
screen "设置画面" 1280x740, template "模板_设置"
   on GenerateScreen: "TitleUpdater"()
   TextField "Text Field_2" at 90,72 size 116x49; Text '总捻度:'
   TextField "Text Field_6" at 320,72 size 107x49; Text '捻/米'
   TextField "Text Field_19" at 674,70 size 140x49; Text '捻缩捻度:'
   TextField "Text Field_20" at 674,133 size 140x49; Text '捻缩距离:'
   TextField "Text Field_21" at 674,196 size 140x49; Text '捻缩时间:'
   TextField "Text Field_22" at 674,259 size 140x49; Text '捻缩速度:'
   TextField "Text Field_15" at 786,14 size 154x42; Text '捻缩设定'
   TextField "Text Field_29" at 753,476 size 140x49; Text '成纱支数:'
   TextField "Text Field_31" at 674,322 size 140x49; Text '卷绕长度:'
   TextField "Text Field_32" at 940,70 size 98x49; Text '捻/米'
   TextField "Text Field_33" at 940,133 size 98x49; Text 'mm'
   TextField "Text Field_34" at 940,196 size 98x49; Text '秒'
   TextField "Text Field_35" at 940,259 size 98x49; Text 'mm/s'
   TextField "Text Field_36" at 940,322 size 98x49; Text 'mm'
   TextField "Text Field_48" at 552,72 size 84x49; Text '秒'
   TextField "Text Field_40" at 791,420 size 228x42; Text '成形、张力设定'
   TextField "Text Field_41" at 753,539 size 140x49; Text '纱穗个数:'
   TextField "Text Field_41#mig1" at 753,602 size 140x49; Text '单纱张力:'
   TextField "Text Field_14" at 142,14 size 336x42; Text '捻度设定分配/锭速设定'
   TextField "Text Field_25" at 96,477 size 133x48; Text '总牵伸:'
   TextField "Text Field_26" at 96,540 size 133x49; Text '送条牵伸:'
   TextField "Text Field_1" at 365,420 size 193x42; Text '牵伸设定分配'
   TextField "Text Field_28" at 348,540 size 212x49; Text '第一牵伸(3段):'
   TextField "Text Field_37" at 348,603 size 212x49; Text '集中牵伸区(3段):'
   TextField "Text Field_38" at 348,477 size 212x48; Text '第一牵伸区(3段):'
   TextField "Text Field_39" at 666,477 size 32x48; Text 'mm'
   TextField "Text Field_42" at 666,603 size 32x49; Text 'mm'
   TextField "Text Field_27" at 43,603 size 186x49; Text '分散牵伸(2段):'
   SymbolicIOField "符号 IO 域_1" at 229,420 size 106x44; TextOn '1'; TextOff '0'; TextList "QainShen_Select"
      ProcessValue <- "ST_HMI_Var_HMI_i16_QianShen_Select"
   IOField "IO Field_14" at 229,477 size 106x48; FormatPattern 9.99
      ProcessValue <- "ST_HMI_Var_HMI_r64QianShen_All"
   IOField "IO Field_15" at 229,540 size 106x49; FormatPattern 9.999
      ProcessValue <- "ST_HMI_Var_HMI_r64QianShen_WuNian"
   IOField "IO Field_17" at 560,540 size 93x49; FormatPattern 9.99
      ProcessValue <- "ST_HMI_Var_HMI_r64QianShen_First"
   IOField "IO Field_20" at 560,603 size 93x49; FormatPattern 99
      ProcessValue <- "ST_HMI_Var_HMI_r64QianShen_finalArea"
   IOField "IO Field_21" at 560,477 size 93x48; FormatPattern 999
      ProcessValue <- "ST_HMI_Var_HMI_r64QianShen_FirstArea"
   IOField "IO Field_16" at 229,603 size 106x49; FormatPattern 9.99
      ProcessValue <- "ST_HMI_Var_HMI_r64QianShen_FenSan"
   TextField "Text Field_3" at 66,136 size 140x47; Text '牵伸捻度:'
   IOField "IO Field_1" at 208,136 size 104x49; FormatPattern 999
      on OnFinishInput: SetBit("ST_Calculation_Var_HMI_bo_Calculation_0_Start"); SetTag("ST_Calculation_Var_g_i16_Calculation_0_3_Select_Status", 1)
      ProcessValue <- "ST_HMI_Var_HMI_r64NianDu_QianShen_Best"
   TextField "Text Field_4" at 320,136 size 107x49; Text '捻/米'
   TextField "Text Field_5" at 552,136 size 84x49; Text '转/分'
   IOField "IO Field_3" at 208,200 size 104x49; FormatPattern 9.99
      on OnFinishInput: SetBit("ST_Calculation_Var_HMI_bo_Calculation_0_Start"); SetTag("ST_Calculation_Var_g_i16_Calculation_0_3_Select_Status", 1)
      ProcessValue <- "ST_HMI_Var_HMI_r64Ratio_PositiveAccel_Jerk_JiaNian"
   TextField "Text Field_8" at 66,264 size 140x47; Text '追捻:'
   Button "OBJECT_107" at 208,264 size 104x48; TextOff '启用 / EXIT'
      on Release: SetBit("ST_HMI_Var_HMI_boNianDu_3")
      on Change: SetBit("ST_Calculation_Var_HMI_bo_Calculation_0_Start"); SetTag("ST_Calculation_Var_g_i16_Calculation_0_3_Select_Status", 1)
      Appearance <- "ST_HMI_Var_HMI_boNianDu_3"
   Button "OBJECT_1" at 432,264 size 112x48; TextOff '停用 / EXIT'
      on Release: ResetBit("ST_HMI_Var_HMI_boNianDu_3")
      on Change: SetBit("ST_Calculation_Var_HMI_bo_Calculation_0_Start"); SetTag("ST_Calculation_Var_g_i16_Calculation_0_3_Select_Status", 1)
      Appearance <- "ST_HMI_Var_HMI_boNianDu_3"
   TextField "Text Field_9" at 24,328 size 182x47; Text '追捻开始捻度:'
   IOField "IO Field_4" at 208,328 size 104x49; FormatPattern 9999
      on OnFinishInput: SetBit("ST_Calculation_Var_HMI_bo_Calculation_0_Start"); SetTag("ST_Calculation_Var_g_i16_Calculation_0_3_Select_Status", 1)
      ProcessValue <- "ST_HMI_Var_HMI_r64NianDu_1"
   TextField "Text Field_10" at 328,328 size 84x49; Text '捻/米'
   TextField "Text Field_11" at 552,328 size 84x49; Text '转/分'
   TextField "Text Field_12" at 320,200 size 107x47; Text '加速度:'
   IOField "IO Field_5" at 432,328 size 112x49; FormatPattern 99999
      on OnFinishInput: SetBit("ST_Calculation_Var_HMI_bo_Calculation_0_Start"); SetTag("ST_Calculation_Var_g_i16_Calculation_0_3_Select_Status", 1)
      ProcessValue <- "ST_HMI_Var_HMI_r64NianSu_2"
   TextField "Text Field_7" at 48,202 size 158x47; Text '加速度比例:'
   IOField "IO Field_43" at 208,72 size 104x49; FormatPattern 9999
      on OnFinishInput: SetBit("ST_Calculation_Var_HMI_bo_Calculation_0_Start"); SetTag("ST_Calculation_Var_g_i16_Calculation_0_3_Select_Status", 1)
      ProcessValue <- "ST_HMI_Var_HMI_r64NianDu_all"
   IOField "IO Field_13" at 432,72 size 112x49; FormatPattern 99.9
      ProcessValue <- "ST_HMI_Var_HMI_r64Time_JiaNian"
      Appearance <- "ST_HMI_Var_HMI_boAlarm_NianDu_Time"
   IOField "IO Field_9" at 814,70 size 112x49; FormatPattern 9999
      on OnFinishInput: SetBit("ST_Calculation_Var_HMI_bo_Calculation_0_Start"); SetTag("ST_Calculation_Var_g_i16_Calculation_0_3_Select_Status", 1)
      ProcessValue <- "ST_HMI_Var_HMI_r64NianDu_NianSuo"
   IOField "IO Field_10" at 814,133 size 112x49; FormatPattern 999
      on OnFinishInput: SetBit("ST_Calculation_Var_HMI_bo_Calculation_0_Start")
      Appearance <- "ST_HMI_Var_HMI_boAlarm_NianSuo_PosNon"
      ProcessValue <- "ST_HMI_Var_HMI_r64Position_NianSuo"
   IOField "IO Field_11" at 814,196 size 112x49; FormatPattern 99.9
      ProcessValue <- "ST_HMI_Var_HMI_r64Time_NianSuo"
   IOField "IO Field_12" at 814,259 size 112x49; FormatPattern 99.9
      ProcessValue <- "ST_HMI_Var_HMI_r64Velocity_NianSuo"
      Appearance <- "ST_HMI_Var_HMI_boAlarm_NianSuo_SuDuOver"
   IOField "IO Field_19" at 814,322 size 112x49; FormatPattern 9999
      ProcessValue <- "ST_HMI_Var_HMI_r64Length_JuanRao"
   IOField "IO Field_18" at 907,476 size 126x49; FormatPattern 99.99
      ProcessValue <- "ST_HMI_Var_HMI_r64ZhiShu_ChengSha"
   IOField "IO Field_75" at 907,539 size 126x49; FormatPattern 9999
      ProcessValue <- "ST_HMI_Var_HMI_r64_ShuLiang_ShaSui"
   IOField "IO Field_76" at 907,602 size 126x49; FormatPattern 999.9
      ProcessValue <- "ST_HMI_Var_HMI_r64_LuoSha_Force_DanSha_ZhangLi_FangKai"
   IOField "IO Field_2" at 432,136 size 112x49; FormatPattern 99999
      ProcessValue <- "ST_HMI_Var_HMI_r64NianSu_Max"
      Appearance <- "ST_HMI_Var_HMI_boAlarm_NianDu_Time"
   IOField "IO Field_6" at 432,200 size 112x49; FormatPattern 99999
      Visibility <- "ST_Calculation_Var_Date_Temp"
      ProcessValue <- "ST_Calculation_Var_g_r64Axis_DingZi_PositiveAccel_Buffer_JiaNian{0}"
      Appearance <- "ST_HMI_Var_HMI_boAlarm_NianDu_Time"
   IOField "IO Field_8" at 432,200 size 112x49; FormatPattern 99999
      Visibility <- "ST_Calculation_Var_Date_Temp"
      ProcessValue <- "ST_Calculation_Var_g_r64Axis_DingZi_PositiveAccel_Buffer_JiaNian{1}"
      Appearance <- "ST_HMI_Var_HMI_boAlarm_NianDu_Time"
   TextField "文本域_5" at 1,304 size 880x170; Text '捻度报警！设置捻度为 ，实际捻度为 ， 已自动停止，请检查设置画面参数，重新设置总捻度， 检查设置其他参数，使画面上的参数没有红色闪烁，然 后按“启动”，若继续出现此报警，请从生头重新开始'
      Visibility <- "ST_HMI_Var_HMI_i16_NianduAlarmStatus"
   IOField "IO Field_7" at 322,305 size 86x32; FormatPattern 9999
      on OnFinishInput: SetBit("ST_Calculation_Var_HMI_bo_Calculation_0_Start"); SetTag("ST_Calculation_Var_g_i16_Calculation_0_3_Select_Status", 1)
      Visibility <- "ST_HMI_Var_HMI_i16_NianduAlarmStatus"
      ProcessValue <- "ST_HMI_Var_HMI_r64NianDu_all"
   IOField "IO Field_22" at 601,305 size 86x32; FormatPattern 9999
      Visibility <- "ST_HMI_Var_HMI_i16_NianduAlarmStatus"
      ProcessValue <- "ST_HMI_Var_HMI_r64Niandu_all_Current"
   Button "按钮_16" at 734,414 size 137x44; TextOff '知道了'
      on Click: SetTag("ST_HMI_Var_HMI_i16_NianduAlarmStatus", 0); SetBit("ST_Calculation_Var_HMI_bo_Calculation_0_Start"); ResetBit("ST_HMI_Var_HMI_bo_XiangLing")
      Visibility <- "ST_HMI_Var_HMI_i16_NianduAlarmStatus"
   Circle "圆_4" at 774,325 size 60x60
      Visibility <- "ST_HMI_Var_HMI_i16_NianduAlarmStatus"
      Appearance <- "ST_HMI_Var_HMI_bo_XiangLing"
   TextField "文本域_10" at 7,311 size 880x170; Text '锭子不转报警！请至报警画面解除报警，然后点击“退 出紧急停止”，点击“启动”开机，或者按正常步骤断电 重启，然后开机'
      Visibility <- "ST_HMI_Var_HMI_i16_Dingzi_50102AlarmStatus"
   Button "按钮_6" at 732,413 size 137x44; TextOff '知道了'
      on Click: SetTag("ST_HMI_Var_HMI_i16_Dingzi_50102AlarmStatus", 0); ResetBit("ST_HMI_Var_HMI_bo_XiangLing")
      Visibility <- "ST_HMI_Var_HMI_i16_Dingzi_50102AlarmStatus"
   Circle "圆_1" at 772,324 size 60x60
      Visibility <- "ST_HMI_Var_HMI_i16_Dingzi_50102AlarmStatus"
      Appearance <- "ST_HMI_Var_HMI_bo_XiangLing"

screen "时间显示" 1280x740, template "模板_根"
   on GenerateScreen: "TitleUpdater"(); "timeConverse"()
   Button "HmiScreenItemData_8" at 1120,65 size 159x47; TextOn '向后'; TextOff '向后'
      on Release: ActivateScreen("友联走架智控系统", 0)
   Button "按钮_1" at 174,88 size 95x82; TextOff '出车'
      Appearance <- "ST_Main_Var_g_i16_Automatic_Status"
   Button "按钮_2" at 321,88 size 95x82; TextOff '加捻'
      Appearance <- "ST_Main_Var_g_i16_Automatic_Status"
   Button "按钮_3" at 467,88 size 96x82; TextOff '退绕'
      Appearance <- "ST_Main_Var_g_i16_Automatic_Status"
   Button "按钮_4" at 614,88 size 95x82; TextOff '进车'
      Appearance <- "ST_Main_Var_g_i16_Automatic_Status"
   Button "按钮_5" at 760,88 size 96x82; TextOff '周期'
      Appearance <- "ST_Main_Var_g_i16_Automatic_Status"
   TextField "文本域_1" at 51,360 size 207x37; Text '系统总运行时间:'
   TextField "文本域_2" at 346,360 size 56x37; Text '年'
   TextField "文本域_4" at 460,360 size 56x37; Text '天'
   TextField "文本域_5" at 563,360 size 56x37; Text '时'
   TextField "文本域_6" at 661,360 size 56x37; Text '分'
   TextField "文本域_7" at 760,360 size 56x37; Text '秒'
   IOField "IO Field_23" at 174,183 size 95x55; FormatPattern 99.99
      ProcessValue <- "ST_Main_Var_g_r64_Time_chuche"
   IOField "IO Field_24" at 321,183 size 95x55; FormatPattern 99.99
      ProcessValue <- "ST_Main_Var_g_r64_Time_jianian"
   IOField "IO Field_25" at 467,183 size 96x55; FormatPattern 99.99
      ProcessValue <- "ST_Main_Var_g_r64_Time_tuirao"
   IOField "IO Field_26" at 614,183 size 95x55; FormatPattern 99.99
      ProcessValue <- "ST_Main_Var_g_r64_Time_juanrao"
   IOField "IO Field_27" at 760,183 size 96x55; FormatPattern 99.99
      ProcessValue <- "ST_Main_Var_g_r64_Time_Once"
   IOField "IO Field_29" at 269,350 size 72x55; FormatPattern 999
      ProcessValue <- "VBS_time_year"
   IOField "IO Field_30" at 385,350 size 68x55; FormatPattern 999
      ProcessValue <- "VBS_time_day"
   IOField "IO Field_30#mig1" at 499,350 size 55x55; FormatPattern 99
      ProcessValue <- "VBS_time_hour"
   IOField "IO Field_31" at 600,350 size 55x55; FormatPattern 99
      ProcessValue <- "VBS_time_min"
   IOField "IO Field_32" at 701,350 size 52x55; FormatPattern 99
      ProcessValue <- "VBS_time_sec"

screen "手动画面" 1280x740, template "模板_动画"
   on GenerateScreen: "TitleUpdater"()
   Button "HmiScreenItemData_2" at 1150,25 size 130x47; TextOn '手动设置'; TextOff '手动设置'
      on Release: ActivateScreen("手动设置", 0)
   Button "OBJECT_106" at 904,14 size 231x33; TextOff '手动 / EXIT'; TextList "mode_enabled_1"
      ProcessValue <- "ST_Main_Var_g_i16_Mode_Enabled"
      Appearance <- "ST_Main_Var_g_i16_Mode_Enabled"
   Button "OBJECT_2" at 172,583 size 119x60; TextOff '启动 / EXIT'
      on Release: ResetBit("ST_HMI_Var_HMI_bo_ZiDong_QiDong")
      on Press: SetBit("ST_HMI_Var_HMI_bo_ZiDong_QiDong")
      Appearance <- "ST_Main_Var_g_i16_Start_Position_Status"
      Visibility <- "ST_Main_Var_g_i16_Mode_Enabled"
   Button "OBJECT_3" at 762,15 size 119x65; TextOff 'SLM / EXIT'
      on Press: SetBit("ST_Main_Var_g_SLM_enable_status")
      Appearance <- "ST_Main_Var_g_SLM_enable_status"
   Button "OBJECT_4" at 9,583 size 119x60; TextOff '急停 / EXIT'
      on Click: InvertBit("ST_Main_Var_g_bo_ZiDong_JiTing")
      Appearance <- "ST_Main_Var_g_bo_ZiDong_JiTing"
   Button "OBJECT_15" at 474,16 size 119x65; TextOff '电源通 / EXIT'
      Appearance <- "PLCAddressVar_g_bo_DI_1_D435_X122_2"
   Button "OBJECT_16" at 619,14 size 119x65; TextOff '电源断 / EXIT'
      on Release: ResetBit("ST_HMI_Var_HMI_bo_DianYuan_Duan")
      on Press: SetBit("ST_HMI_Var_HMI_bo_DianYuan_Duan")
   IOField "IO 域_20" at 903,47 size 231x33; Authorization "User administration"; FormatPattern 9
      on Activate: function_f41c6f6c("变量_1")
      ProcessValue <- "ST_Main_Var_g_i16_Manual_Status"
   Button "OBJECT_5" at 172,493 size 119x60; TextOff '手 动 / EXIT'
      on Release: ResetBit("ST_HMI_Var_HMI_bo_Manual")
      on Press: SetBit("ST_HMI_Var_HMI_bo_Manual")
      Appearance <- "ST_Main_Var_g_i16_Manual_Status"
   Button "OBJECT_6" at 9,493 size 119x60; TextOff '去使能 / EXIT'
      on Release: ResetBit("ST_HMI_Var_HMI_bo_Disable")
      on Press: SetBit("ST_HMI_Var_HMI_bo_Disable")
      Appearance <- "ST_Main_Var_g_i16_Disable_Status"
   Button "OBJECT_110" at 335,583 size 119x60; TextOff '停 止 / EXIT'
      on Release: ResetBit("ST_HMI_Var_HMI_bo_ZiDong_TingZhi")
      on Press: SetBit("ST_HMI_Var_HMI_bo_ZiDong_TingZhi")
      Appearance <- "ST_Main_Var_g_i16_Start_Position_Status"
      Visibility <- "ST_Main_Var_g_i16_Mode_Enabled"
   Button "OBJECT_7" at 335,493 size 119x60; TextOff '回起点 / EXIT'
      on Release: ResetBit("ST_HMI_Var_HMI_bo_Start_Position")
      on Press: SetBit("ST_HMI_Var_HMI_bo_Start_Position")
      Appearance <- "ST_Main_Var_g_i16_Mode_Enabled"
   Group "Group_手动按钮" at 496,493 size 760x150
   Button "OBJECT_17" at 496,493 size 120x60; TextOff '出车 / EXIT'
      on Release: ResetBit("ST_HMI_Var_HMI_bo_ChuChe")
      on Press: SetBit("ST_HMI_Var_HMI_bo_ChuChe")
      Appearance <- "ST_HMI_Var_HMI_bo_ChuChe"
      Visibility <- "ST_Main_Var_g_i16_Mode_Enabled"
   Button "OBJECT_18" at 656,493 size 120x60; TextOff '送条 / EXIT'
      on Release: InvertBit("ST_HMI_Var_HMI_bo_SongTiao")
      Appearance <- "ST_HMI_Var_HMI_bo_SongTiao"
      Visibility <- "ST_Main_Var_g_i16_Mode_Enabled"
   Button "OBJECT_19" at 816,493 size 120x60; TextOff '退绕 / EXIT'
      on Release: ResetBit("ST_HMI_Var_HMI_bo_TuiRao")
      on Press: SetBit("ST_HMI_Var_HMI_bo_TuiRao")
      Appearance <- "ST_HMI_Var_HMI_bo_TuiRao"
      Visibility <- "ST_Main_Var_g_i16_Mode_Enabled"
   Button "OBJECT_20" at 976,493 size 120x60; TextOff '成形弓降 / EXIT'
      on Release: ResetBit("ST_HMI_Var_HMI_bo_ChengXing_Down")
      on Press: SetBit("ST_HMI_Var_HMI_bo_ChengXing_Down")
      Appearance <- "ST_HMI_Var_HMI_bo_ChengXing_Down"
      Visibility <- "ST_Main_Var_g_i16_Mode_Enabled"
   Button "OBJECT_21" at 1136,493 size 120x60; TextOff '张力弓升 / EXIT'
      on Release: ResetBit("ST_HMI_Var_HMI_bo_ZhangLi_Up")
      on Press: SetBit("ST_HMI_Var_HMI_bo_ZhangLi_Up")
      Appearance <- "ST_HMI_Var_HMI_bo_ZhangLi_Up"
      Visibility <- "ST_Main_Var_g_i16_Mode_Enabled"
   Button "OBJECT_22" at 496,583 size 120x60; TextOff '进车 / EXIT'
      on Release: ResetBit("ST_HMI_Var_HMI_bo_JinChe")
      on Press: SetBit("ST_HMI_Var_HMI_bo_JinChe")
      Appearance <- "ST_HMI_Var_HMI_bo_JinChe"
      Visibility <- "ST_Main_Var_g_i16_Mode_Enabled"
   Button "OBJECT_23" at 656,583 size 120x60; TextOff '加捻 / EXIT'
      on Release: ResetBit("ST_HMI_Var_HMI_bo_JiaNian")
      on Press: SetBit("ST_HMI_Var_HMI_bo_JiaNian")
      Appearance <- "ST_Main_Var_g_bo_JianNian_Jog_Status"
      Visibility <- "ST_Main_Var_g_i16_Mode_Enabled"
   Button "OBJECT_24" at 816,583 size 120x60; TextOff '卷绕 / EXIT'
      on Release: ResetBit("ST_HMI_Var_HMI_bo_JuanRao")
      on Press: SetBit("ST_HMI_Var_HMI_bo_JuanRao")
      Appearance <- "ST_HMI_Var_HMI_bo_JuanRao"
      Visibility <- "ST_Main_Var_g_i16_Mode_Enabled"
   Button "OBJECT_25" at 976,583 size 120x60; TextOff '成形弓升 / EXIT'
      on Release: ResetBit("ST_HMI_Var_HMI_bo_ChengXing_Up")
      on Press: SetBit("ST_HMI_Var_HMI_bo_ChengXing_Up")
      Appearance <- "ST_HMI_Var_HMI_bo_ChengXing_Up"
      Visibility <- "ST_Main_Var_g_i16_Mode_Enabled"
   Button "OBJECT_26" at 1136,583 size 120x60; TextOff '张力弓降 / EXIT'
      on Release: ResetBit("ST_HMI_Var_HMI_bo_ZhangLi_Down")
      on Press: SetBit("ST_HMI_Var_HMI_bo_ZhangLi_Down")
      Appearance <- "ST_HMI_Var_HMI_bo_ZhangLi_Down"
      Visibility <- "ST_Main_Var_g_i16_Mode_Enabled"

screen "手动设置" 1280x740, template "模板_根"
   on GenerateScreen: "TitleUpdater"()
   Button "HmiScreenItemData_3" at 1119,125 size 159x47; TextOn '向后'; TextOff '向后'
      on Release: ActivateScreen("手动画面", 0)
   IOField "IO 域_20" at 80,185 size 120x41; FormatPattern 99999999
      on Activate: function_f41c6f6c("变量_1")
      ProcessValue <- "ST_HMI_Var_HMI_r64Velocity_Jog_Chuche"
   TextField "文本域_19" at 886,57 size 172x38; Text '当前登录用户'
   IOField "IO 域_15" at 914,98 size 122x41; FormatPattern ?????????????
      ProcessValue <- "user_name"
   IOField "IO 域_2" at 80,417 size 120x41; FormatPattern 99999999
      ProcessValue <- "ST_HMI_Var_HMI_r64Velocity_Jog_JinChe"
   IOField "IO 域_3" at 232,417 size 120x41; FormatPattern 999999999
      ProcessValue <- "ST_HMI_Var_HMI_r64Velocity_Jog_JiaNian"
   IOField "IO 域_5" at 384,417 size 120x41; FormatPattern 999999999
      ProcessValue <- "ST_HMI_Var_HMI_r64Velocity_Jog_JuanRao"
   IOField "IO 域_4" at 232,185 size 120x41; FormatPattern 99999999
      ProcessValue <- "ST_HMI_Var_HMI_r64Velocity_Jog_SongTiao"
   IOField "IO 域_16" at 384,185 size 120x41; FormatPattern 999999999
      ProcessValue <- "ST_HMI_Var_HMI_r64Velocity_Jog_TuiRao"
   IOField "IO 域_6" at 536,416 size 120x41; Authorization "User administration"; FormatPattern 99999999
      ProcessValue <- "ST_HMI_Var_HMI_r64Velocity_Jog_ChengXing_Up"
   IOField "IO 域_7" at 536,186 size 120x41; Authorization "User administration"; FormatPattern 99999999
      ProcessValue <- "ST_HMI_Var_HMI_r64Velocity_Jog_ChengXing_Down"
   IOField "IO 域_9" at 688,184 size 120x41; Authorization "User administration"; FormatPattern 99999999
      ProcessValue <- "ST_HMI_Var_HMI_r64Velocity_Jog_ZhangLi_Up"
   IOField "IO 域_10" at 688,416 size 120x41; Authorization "User administration"; FormatPattern 99999999
      ProcessValue <- "ST_HMI_Var_HMI_r64Velocity_Jog_ZhangLi_Down"
   IOField "IO 域_21" at 80,253 size 120x41; FormatPattern 99999999
      on Activate: function_f41c6f6c("变量_1")
      ProcessValue <- "ST_HMI_Var_HMI_r64AccVelocity_Jog_ChuChe"
   IOField "IO 域_8" at 80,485 size 120x41; FormatPattern 99999999
      ProcessValue <- "ST_HMI_Var_HMI_r64AccVelocity_Jog_JinChe"
   Button "OBJECT_119" at 328,588 size 177x68; TextOff '选择市电模式 / EXIT'; Authorization "Operate_5"
      on Press: SetBit("ST_HMI_Var_HMI_Bo_Feed_On_Off_Select")
      Appearance <- "ST_HMI_Var_HMI_Bo_Feed_On_Off_Select"
   Button "OBJECT_120" at 579,588 size 177x68; TextOff '选择发电模式 / EXIT'; Authorization "Operate_5"
      on Press: ResetBit("ST_HMI_Var_HMI_Bo_Feed_On_Off_Select")
      Appearance <- "ST_HMI_Var_HMI_Bo_Feed_On_Off_Select"
   Button "OBJECT_5" at 80,80 size 120x80; TextOff '出车 / EXIT'
      on Release: ResetBit("ST_HMI_Var_HMI_bo_ChuChe")
      on Press: SetBit("ST_HMI_Var_HMI_bo_ChuChe")
      Appearance <- "ST_HMI_Var_HMI_bo_ChuChe"
   Button "OBJECT_7" at 232,80 size 120x80; TextOff '送条 / EXIT'
      on Release: InvertBit("ST_HMI_Var_HMI_bo_SongTiao")
      Appearance <- "ST_HMI_Var_HMI_bo_SongTiao"
   Button "OBJECT_9" at 384,80 size 120x80; TextOff '退绕 / EXIT'
      on Release: ResetBit("ST_HMI_Var_HMI_bo_TuiRao")
      on Press: SetBit("ST_HMI_Var_HMI_bo_TuiRao")
      Appearance <- "ST_HMI_Var_HMI_bo_TuiRao"
   Button "OBJECT_12" at 536,80 size 120x80; TextOff '成形弓降 / EXIT'
      on Release: ResetBit("ST_HMI_Var_HMI_bo_ChengXing_Down")
      on Press: SetBit("ST_HMI_Var_HMI_bo_ChengXing_Down")
      Appearance <- "ST_HMI_Var_HMI_bo_ChengXing_Down"
   Button "OBJECT_13" at 688,80 size 120x80; TextOff '张力弓升 / EXIT'
      on Release: ResetBit("ST_HMI_Var_HMI_bo_ZhangLi_Up")
      on Press: SetBit("ST_HMI_Var_HMI_bo_ZhangLi_Up")
      Appearance <- "ST_HMI_Var_HMI_bo_ZhangLi_Up"
   Button "OBJECT_6" at 81,312 size 120x80; TextOff '进车 / EXIT'
      on Release: ResetBit("ST_HMI_Var_HMI_bo_JinChe")
      on Press: SetBit("ST_HMI_Var_HMI_bo_JinChe")
      Appearance <- "ST_HMI_Var_HMI_bo_JinChe"
   Button "OBJECT_8" at 232,312 size 120x80; TextOff '加捻 / EXIT'
      on Release: ResetBit("ST_HMI_Var_HMI_bo_JiaNian")
      on Press: SetBit("ST_HMI_Var_HMI_bo_JiaNian")
      Appearance <- "ST_Main_Var_g_bo_JianNian_Jog_Status"
   Button "OBJECT_10" at 384,312 size 120x80; TextOff '卷绕 / EXIT'
      on Release: ResetBit("ST_HMI_Var_HMI_bo_JuanRao")
      on Press: SetBit("ST_HMI_Var_HMI_bo_JuanRao")
      Appearance <- "ST_HMI_Var_HMI_bo_JuanRao"
   Button "OBJECT_11" at 536,312 size 120x80; TextOff '成形弓升 / EXIT'
      on Release: ResetBit("ST_HMI_Var_HMI_bo_ChengXing_Up")
      on Press: SetBit("ST_HMI_Var_HMI_bo_ChengXing_Up")
      Appearance <- "ST_HMI_Var_HMI_bo_ChengXing_Up"
   Button "OBJECT_14" at 688,312 size 120x80; TextOff '张力弓降 / EXIT'
      on Release: ResetBit("ST_HMI_Var_HMI_bo_ZhangLi_Down")
      on Press: SetBit("ST_HMI_Var_HMI_bo_ZhangLi_Down")
      Appearance <- "ST_HMI_Var_HMI_bo_ZhangLi_Down"
   Button "OBJECT_1" at 536,482 size 120x80; TextOff '成形弓 抱闸松开 EXIT'
      on Press: InvertBit("ST_HMI_Var_HMI_bo_ChengXing_Holding_Brake_Open")
      Appearance <- "ST_HMI_Var_HMI_bo_ChengXing_Holding_Brake_Open"
      Visibility <- "ST_Main_Var_g_i16_Mode_Enabled"
      ObjectEnable <- "ST_Main_Var_g_i16_Disable_Status"
   Button "OBJECT_2" at 688,482 size 120x80; TextOff '张力弓 抱闸松开 EXIT'
      on Press: InvertBit("ST_HMI_Var_HMI_bo_ZhangLi_Holding_Brake_Open")
      Appearance <- "ST_HMI_Var_HMI_bo_ZhangLi_Holding_Brake_Open"
      Visibility <- "ST_Main_Var_g_i16_Mode_Enabled"
      ObjectEnable <- "ST_Main_Var_g_i16_Disable_Status"
   Button "OBJECT_3" at 385,482 size 120x80; TextOff '走车 抱闸松开 EXIT'
      on Press: InvertBit("ST_HMI_Var_HMI_bo_ZouChe_Holding_Brake_Open")
      Visibility <- "ST_Main_Var_g_i16_Mode_Enabled"
      ObjectEnable <- "ST_Main_Var_g_i16_Disable_Status"
      Appearance <- "ST_HMI_Var_HMI_bo_ZouChe_Holding_Brake_Open"

screen "调试画面" 1280x740, template "模板_调试"
   on GenerateScreen: "TitleUpdater"()
   TextField "Text Field_44" at 273,417 size 327x41; Text '退绕曲线拐点比例 / パッキングオフ湾曲点比例 / 언와인딩 곡선 변곡점 비율'
   TextField "Text Field_46" at 273,468 size 327x41; Text '退绕圈数比例 / パッキングオフ巻取比例 / 언와인딩 랩수 비율'
   TextField "Text Field_37" at 276,210 size 327x41; Text '卷绕速度中点调整值—初始值 / 中間点の取り巻き速度調整値ー初期値 / 와인딩 속도 중심점조정값-초기값'
   TextField "Text Field_38" at 276,261 size 327x41; Text '卷绕速度末点调整值—初始值 / 終了時点の取り巻き速度調整値ー初期値 / 와인딩 속도 종료점조정값-초기값'
   TextField "Text Field_39" at 276,159 size 327x41; Text '卷绕张力弓目标值—满纱时 / カウンターフォーラーの目標値ー満巻時 / 와인딩 장력 호랑 목표값-만사일시'
   TextField "Text Field_40" at 276,108 size 327x41; Text '卷绕张力弓目标值—最大直径时 / カウンターフォーラーの目標値ー最大直径時 / 와이딩 장력 호랑목표값-최대직경일시'
   TextField "Text Field_41" at 276,57 size 327x41; Text '卷绕张力弓目标值—生头时 / カウンターフォーラーの目標値ー巻始め / 와인딩 장력호랑 목표값-실시작점'
   TextField "Text Field_45" at 276,312 size 327x41; Text '卷绕张力弓反馈增益 / カウンターフォーラーのフィードバック増幅 / 와인딩 장력호랑 피드백 게인'
   TextField "Text Field_1" at 276,561 size 327x41; Text '存绕锭子加速度 / 逆巻取スピンドル加速度 / 와인딩 스핀들 가속'
   TextField "Text Field_42" at 276,614 size 327x41; Text '存绕锭子速度比例 / 逆巻取スピンドル回転速度比例 / 와인딩 스핀들 속도 비율'
   TextField "Text Field_14" at 154,2 size 233x42; Text '卷绕相关 / 巻取関係 / 와인딩 관련'
   TextField "Text Field_3" at 153,365 size 233x42; Text '退绕相关 / パッキングオフ関連 / 언와인딩 관련'
   TextField "Text Field_4" at 153,518 size 233x42; Text '存绕相关 / 逆巻取関連 / 와인딩관련'
   TextField "Text Field_5" at 658,2 size 233x42; Text '其他 / その他 / 기타'
   IOField "IO Field_4" at 658,429 size 112x42; FormatPattern 9.99
      on OnFinishInput: SetBit("ST_Calculation_Var_HMI_bo_Calculation_0_Start"); SetTag("ST_Calculation_Var_g_i16_Calculation_0_3_Select_Status", 1)
      ProcessValue <- "ST_TO_DZ_FU_Var_HMI_r64Ratio_PositiveAccelStartJerk_JiaNian"
   IOField "IO Field_6" at 658,483 size 112x42; FormatPattern 9.99
      on OnFinishInput: SetBit("ST_Calculation_Var_HMI_bo_Calculation_0_Start"); SetTag("ST_Calculation_Var_g_i16_Calculation_0_3_Select_Status", 1)
      ProcessValue <- "ST_TO_DZ_FU_Var_HMI_r64Ratio_PositiveAccelEndJerk_JiaNian"
   IOField "IO Field_9" at 658,537 size 112x42; FormatPattern 99.99
      ProcessValue <- "ST_HMI_Var_HMI_r64_DingZi_Zouche_ratio_KongDing_65_1"
   IOField "IO Field_5" at 658,322 size 112x42; FormatPattern 9.99
      on OnFinishInput: SetBit("ST_Calculation_Var_HMI_bo_Calculation_0_Start"); SetTag("ST_Calculation_Var_g_i16_Calculation_0_3_Select_Status", 1)
      ProcessValue <- "ST_HMI_Var_HMI_r64Ratio_PositiveAccel_Jerk_JiaNian"
   TextField "Text Field_58" at 791,163 size 230x41; Text '生头中间停止位置 / 自動停止位置 / 스레딩중 정지위치'
   TextField "Text Field_8" at 791,56 size 230x41; Text '毛轴头数 / 篠棒本数 / 시누 세부샤프트개수'
   TextField "Text Field_2" at 791,109 size 230x41; Text '生头起点位置 / 口付け開始点位置 / 스레딩시작점 위치'
   TextField "Text Field_6" at 790,216 size 230x41; Text '自动停止位置 / 自動停止位置 / 자동정지위치'
   TextField "Text Field_7" at 790,270 size 230x41; Text '出车停止位置 / 自動停止位置 / 외진정지위치'
   TextField "Text Field_12" at 790,377 size 230x41; Text '锭子加速度'
   TextField "Text Field_9" at 790,430 size 230x41; Text '锭子+Jerk比例'
   TextField "Text Field_11" at 790,484 size 230x41; Text '锭子-Jerk比例'
   TextField "Text Field_13" at 790,538 size 230x41; Text '光锭卷绕传动比1'
   TextField "Text Field_10" at 790,323 size 230x41; Text '锭子加速度比例 / 自動停止位置 / 외진정지위치'
   IOField "IO Field_38" at 658,162 size 112x42; FormatPattern 999
      ProcessValue <- "ST_HMI_Var_HMI_r64Axis_ZouChe_Position_KongDing_12"
   IOField "IO Field_41" at 658,55 size 112x42; FormatPattern 99
      ProcessValue <- "ST_HMI_Var_HMI_r64_MaoZhou_TouShu"
   IOField "IO Field_10" at 658,108 size 112x42; FormatPattern 999.9
      ProcessValue <- "ST_HMI_Var_HMI_r64Axis_ZouChe_Position_ShengTou_Start_Position"
   IOField "IO Field_28" at 154,312 size 108x40; FormatPattern 99.99
      ProcessValue <- "ST_HMI_Var_HMI_r64_k_ZhangLi_Rate"
   IOField "IO Field_21" at 154,260 size 108x41; FormatPattern 99.99
      ProcessValue <- "ST_HMI_Var_HMI_g1_n_delt_new_0"
   IOField "IO Field_20" at 154,208 size 108x41; FormatPattern 99.99
      ProcessValue <- "ST_HMI_Var_HMI_f1_n_delt_new_0"
   IOField "IO Field_22" at 154,157 size 108x40; FormatPattern 99.99
      ProcessValue <- "ST_HMI_Var_HMI_r64Axis_1_ZhangLi_Position_JuanRao_Set_N"
   IOField "IO Field_23" at 154,106 size 108x40; FormatPattern 99.99
      ProcessValue <- "ST_HMI_Var_HMI_r64Axis_1_ZhangLi_Position_JuanRao_Set_ND"
   IOField "IO Field_24" at 154,55 size 108x40; FormatPattern 99.99
      ProcessValue <- "ST_HMI_Var_HMI_r64Axis_1_ZhangLi_Position_JuanRao_Set_0"
   IOField "IO Field_57" at 154,417 size 109x41; FormatPattern 9.99
      ProcessValue <- "ST_HMI_Var_HMI_k_TuiRao"
   IOField "IO Field_58" at 154,468 size 109x41; FormatPattern 9.99
      ProcessValue <- "ST_HMI_Var_HMI_scalevalue_Cam_3"
   IOField "IO Field_1" at 154,572 size 108x40; FormatPattern 99999
      ProcessValue <- "ST_Main_Var_g_r64Axis_DingZi_PositiveAccel_CunRao"
   IOField "IO Field_25" at 154,625 size 108x40; FormatPattern 99.99
      ProcessValue <- "ST_Main_Var_g_r64Axis_DingZi_Velocity_CunRao_ratio"
   IOField "IO Field_2" at 658,215 size 112x42; FormatPattern 99.9
      ProcessValue <- "ST_HMI_Var_HMI_r64Axis_ZouChe_Position_ZiDongTingZhi"
   IOField "IO Field_3" at 658,269 size 112x42; FormatPattern 999
      ProcessValue <- "ST_HMI_Var_HMI_r64Axis_ZouChe_Position_ChuChe_Middle"
   IOField "IO Field_8" at 658,376 size 112x42; FormatPattern 99999
      Visibility <- "ST_Calculation_Var_Date_Temp"
      ProcessValue <- "ST_Calculation_Var_g_r64Axis_DingZi_PositiveAccel_Buffer_JiaNian{1}"
      Appearance <- "ST_HMI_Var_HMI_boAlarm_NianDu_Time"
   IOField "IO Field_7" at 658,376 size 112x42; FormatPattern 99999
      Visibility <- "ST_Calculation_Var_Date_Temp"
      ProcessValue <- "ST_Calculation_Var_g_r64Axis_DingZi_PositiveAccel_Buffer_JiaNian{0}"
      Appearance <- "ST_HMI_Var_HMI_boAlarm_NianDu_Time"

screen "退绕设定" 1280x740, template "模板_设置"
   on GenerateScreen: "TitleUpdater"()
   TextField "Text Field_81" at 292,64 size 196x42; Text '退绕设定'
   TextField "Text Field_82" at 194,134 size 210x56; Text '成形弓速度:'
   TextField "Text Field_84" at 194,208 size 210x56; Text '成形弓加速度:'
   IOField "IO Field_46" at 418,138 size 140x56; FormatPattern 9999
      ProcessValue <- "ST_HMI_Var_HMI_r64Axis_ChengXing_Velocity_TuiRao"
   IOField "IO Field_47" at 418,211 size 140x56; FormatPattern 9999
      ProcessValue <- "ST_HMI_Var_HMI_r64Axis_ChengXing_PositiveAccel_TuiRao"

screen "用户管理" 1280x740, template "模板_根"
   on GenerateScreen: "TitleUpdater"()
   UserView "HmiScreenItemData_7" at 0,0 size 1000x680
   Button "Button_1" at 1055,74 size 170x60; TextOff '登录用户'
      on Press: function_a2a04561()
   Button "Button_2" at 1055,198 size 170x60; TextOff '注销用户'
      on Press: function_f23ef4c9()

screen "13原点设定" 1280x740, template "模板_调试"
   on GenerateScreen: "TitleUpdater"()
   IOField "I/O 域_1" at 996,197 size 88x48; FormatPattern 99
      ProcessValue <- "ST_HMI_Var_HMI_r64StartPosition_Axis_ZouChe_0"
   TextField "文本域_1" at 200,207 size 167x25; Text '走车编码器当前位置'
   IOField "I/O 域_2" at 380,195 size 88x48; FormatPattern 99999
      ProcessValue <- "Axis_ZouChe_positioningState_actualPosition"
   Button "按钮_4" at 868,196 size 76x47; TextOff '出车'
      on Release: ResetBit("ST_HMI_Var_HMI_bo_ChuChe")
      on Press: SetBit("ST_HMI_Var_HMI_bo_ChuChe")
   Button "按钮_5" at 521,195 size 76x47; TextOff '进车'
      on Release: ResetBit("ST_HMI_Var_HMI_bo_JinChe")
      on Press: SetBit("ST_HMI_Var_HMI_bo_JinChe")
   IOField "I/O 域_3" at 996,305 size 88x48; FormatPattern 99.999
      ProcessValue <- "ST_HMI_Var_HMI_r64StartPosition_Axis_1_ZhangLi_0"
   IOField "I/O 域_4" at 996,414 size 88x48
      ProcessValue <- "ST_HMI_Var_HMI_r64StartPosition_Axis_ChengXing_0"
   TextField "文本域_2" at 202,315 size 167x25; Text '张力编码器当前位置'
   IOField "I/O 域_5" at 382,303 size 88x48
      ProcessValue <- "Axis_1_ZhangLi_positioningState_actualPosition"
   Button "按钮_1" at 868,304 size 76x47; TextOff '升'
      on Release: ResetBit("ST_HMI_Var_HMI_bo_ZhangLi_Up")
      on Press: SetBit("ST_HMI_Var_HMI_bo_ZhangLi_Up")
   Button "按钮_2" at 523,303 size 76x47; TextOff '降'
      on Release: ResetBit("ST_HMI_Var_HMI_bo_ZhangLi_Down")
      on Press: SetBit("ST_HMI_Var_HMI_bo_ZhangLi_Down")
   TextField "文本域_3" at 204,425 size 167x25; Text '成形编码器当前位置'
   IOField "I/O 域_6" at 384,413 size 88x48; FormatPattern 999.99
      ProcessValue <- "Axis_ChengXing_positioningState_actualPosition"
   Button "按钮_3" at 523,414 size 76x47; TextOff '升'
      on Release: ResetBit("ST_HMI_Var_HMI_bo_ChengXing_Up")
      on Press: SetBit("ST_HMI_Var_HMI_bo_ChengXing_Up")
   Button "按钮_6" at 868,415 size 76x47; TextOff '降'
      on Release: ResetBit("ST_HMI_Var_HMI_bo_ChengXing_Down")
      on Press: SetBit("ST_HMI_Var_HMI_bo_ChengXing_Down")
   Bar "棒图_1" at 621,196 size 216x49; MaximumValue 90
      ProcessValue <- "Axis_ZouChe_positioningState_actualPosition"
   Bar "棒图_2" at 621,302 size 216x49; MinimumValue 57; MaximumValue 66
      ProcessValue <- "Axis_1_ZhangLi_positioningState_actualPosition"
   Bar "棒图_3" at 621,411 size 216x49; MinimumValue 322; MaximumValue 334
      ProcessValue <- "Axis_ChengXing_positioningState_actualPosition"
   Button "按钮_7" at 200,590 size 163x50; TextOn '微调模式'; TextOff '按下进入微调模式'
      on Release: ResetBit("ST_HMI_Var_HMI_boMinorAdjustment_select")
      on Press: SetBit("ST_HMI_Var_HMI_boMinorAdjustment_select")
   Button "OBJECT_106" at 705,10 size 238x42; TextOff '手动 / EXIT'; TextList "mode_enabled_1"
      ProcessValue <- "ST_Main_Var_g_i16_Mode_Enabled"
      Appearance <- "ST_Main_Var_g_i16_Mode_Enabled"
   TextField "文本域_6" at 297,80 size 791x75; Text '注意： 不要随意修改此页的数据，不当的数据可能导致行程超限撞车的危险！'
   GraphicView "图形视图_2" at 200,71 size 102x99; Picture "图形_2"

screen "14纱管参数" 1280x740, template "模板_调试"
   on GenerateScreen: "TitleUpdater"()
   IOField "IO Field_41" at 148,59 size 112x42; FormatPattern 99.99
      ProcessValue <- "ST_HMI_Var_HMI_r64_h0_s"
   IOField "IO Field_46" at 148,169 size 112x42; FormatPattern 99.99
      ProcessValue <- "ST_HMI_Var_HMI_r64Diameter_ShaGuan_Middle"
   IOField "IO Field_1" at 148,113 size 112x42; FormatPattern 99.99
      ProcessValue <- "ST_HMI_Var_HMI_r64Diameter_ShaGuan_Bottom"
   IOField "IO Field_2" at 148,279 size 112x42
      ProcessValue <- "ST_HMI_Var_HMI_r64Height_ShaGuan_Middle"
   IOField "IO Field_3" at 148,335 size 112x42
      ProcessValue <- "ST_HMI_Var_HMI_r64Height_ShaGuan_Top"
   IOField "IO Field_6" at 148,223 size 112x42; FormatPattern 99.99
      ProcessValue <- "ST_HMI_Var_HMI_r64Diameter_ShaGuan_Top"
   IOField "IO Field_4" at 148,392 size 112x42; FormatPattern 99.9
      ProcessValue <- "ST_HMI_Var_HMI_r64_DingZi_Zouche_ratio_KongDing_9_Shaguan1"
   IOField "IO Field_5" at 640,59 size 112x42; FormatPattern 99.99
      ProcessValue <- "ST_HMI_Var_HMI_r64_h0_s_2"
   IOField "IO Field_7" at 640,169 size 112x42; FormatPattern 99.99
      ProcessValue <- "ST_HMI_Var_HMI_r64Diameter_ShaGuan_Middle_2"
   IOField "IO Field_8" at 640,113 size 112x42; FormatPattern 99.99
      ProcessValue <- "ST_HMI_Var_HMI_r64Diameter_ShaGuan_Bottom_2"
   IOField "IO Field_9" at 640,279 size 112x42
      ProcessValue <- "ST_HMI_Var_HMI_r64Height_ShaGuan_Middle_2"
   IOField "IO Field_10" at 640,335 size 112x42
      ProcessValue <- "ST_HMI_Var_HMI_r64Height_ShaGuan_Top_2"
   IOField "IO Field_11" at 640,223 size 112x42; FormatPattern 99.99
      ProcessValue <- "ST_HMI_Var_HMI_r64Diameter_ShaGuan_Top_2"
   IOField "IO Field_12" at 640,392 size 112x42; FormatPattern 99.9
      ProcessValue <- "ST_HMI_Var_HMI_r64_DingZi_Zouche_ratio_KongDing_9_Shaguan2"
   TextField "Text Field_8" at 286,59 size 332x42; Text '纱管安装高度'
   TextField "Text Field_9" at 286,113 size 332x42; Text '纱管底部直径'
   TextField "Text Field_10" at 286,169 size 332x42; Text '纱管中间直径'
   TextField "Text Field_11" at 286,223 size 332x42; Text '纱管顶部有效直径'
   TextField "Text Field_12" at 286,279 size 332x42; Text '纱管从底部到中间的高度'
   TextField "Text Field_13" at 286,335 size 332x42; Text '纱管从中间到顶部的高度'
   TextField "Text Field_2" at 143,8 size 140x37; Text '标准纱管1:'
   TextField "Text Field_1" at 286,392 size 332x42; Text '空锭-锭子走车传动比'
   TextField "Text Field_3" at 778,59 size 332x42; Text '纱管安装高度'
   TextField "Text Field_4" at 778,113 size 332x42; Text '纱管底部直径'
   TextField "Text Field_5" at 778,169 size 332x42; Text '纱管中间直径'
   TextField "Text Field_6" at 778,223 size 332x42; Text '纱管顶部有效直径'
   TextField "Text Field_7" at 778,279 size 332x42; Text '纱管从底部到中间的高度'
   TextField "Text Field_14" at 778,335 size 332x42; Text '纱管从中间到顶部的高度'
   TextField "Text Field_15" at 635,8 size 140x37; Text '标准纱管2:'
   TextField "Text Field_16" at 778,392 size 332x42; Text '空锭-锭子走车传动比'

screen "牵伸调整画面" 1280x740, template "模板_设置"
   IOField "I/O 域_2" at 378,332 size 106x48; FormatPattern 9.999
      ProcessValue <- "ST_HMI_Var_HMI_r64_QianShen_Add1"
   TextField "Text Field_25" at 85,332 size 296x48; Text '牵伸第一次增加量q1：'
   IOField "I/O 域_1" at 378,414 size 106x48; FormatPattern 9.999
      ProcessValue <- "ST_HMI_Var_HMI_r64_QianShen_Add2"
   TextField "Text Field_1" at 85,414 size 296x48; Text '牵伸第二次增加量q2：'
   IOField "I/O 域_3" at 378,496 size 106x48; FormatPattern 9999
      ProcessValue <- "ST_HMI_Var_HMI_r64_ShaXian_L1"
   TextField "Text Field_2" at 58,496 size 323x48; Text '牵伸第一次增加时纱线米数L1：'
   IOField "I/O 域_4" at 378,578 size 106x48; FormatPattern 9999
      ProcessValue <- "ST_HMI_Var_HMI_r64_ShaXian_L2"
   TextField "Text Field_3" at 66,578 size 315x48; Text '牵伸第二次增加时纱线米数L2：'
   TextField "Text Field_5" at 252,47 size 296x48; Text '牵伸第一次增加量q1：'
   TextField "Text Field_6" at 599,16 size 296x48; Text '牵伸第二次增加量q2：'
   TextField "Text Field_7" at 29,4 size 122x48; Text '总牵伸'
   TextField "Text Field_8" at 984,207 size 122x48; Text '纱线米数'
   TextField "Text Field_9" at 176,259 size 323x48; Text '牵伸第一次增加时纱线米数L1'
   TextField "Text Field_10" at 518,259 size 303x48; Text '牵伸第二次增加时纱线米数L2'
   TextField "Text Field_11" at 904,259 size 149x48; Text '总纱线米数L3'
   IOField "I/O 域_6" at 997,496 size 106x48; FormatPattern 9.999
      ProcessValue <- "ST_HMI_Var_HMI_r64QianShen_All_real"
   TextField "Text Field_12" at 759,496 size 241x48; Text '实时总牵伸：'
   IOField "I/O 域_7" at 997,332 size 106x48; FormatPattern 9.999
      ProcessValue <- "ST_HMI_Var_HMI_r64QianShen_All"
   TextField "Text Field_13" at 759,332 size 241x48; Text '设置的总牵伸：'
   IOField "I/O 域_8" at 997,414 size 106x48; FormatPattern 9.999
      ProcessValue <- "ST_HMI_Var_HMI_r64QianShen_All_object"
   TextField "Text Field_14" at 759,414 size 241x48; Text '调整后的目标总牵伸：'
   IOField "I/O 域_9" at 600,496 size 106x48; FormatPattern 99
      ProcessValue <- "ST_HMI_Var_HMI_r64_Ratio1"
   IOField "I/O 域_10" at 600,578 size 106x48; FormatPattern 99
      ProcessValue <- "ST_HMI_Var_HMI_r64_Ratio2"
   TextField "Text Field_15" at 482,496 size 119x48; Text '百分比1：'
   TextField "Text Field_16" at 485,578 size 119x48; Text '百分比2：'
   TextField "Text Field_4" at 712,496 size 29x48; Text '%'
   TextField "Text Field_17" at 712,578 size 29x48; Text '%'

screen "友联走架智控系统" 1280x740, template "模板_动画"
   on GenerateScreen: "TitleUpdater"(); SetTag("Picture", 1)
   TextField "Text Field_1" at 709,4 size 94x42; Text '满纱周期 / CarriageVelo / キャレージ速度 / 코프완성주기'
   IOField "IO Field_423" at 709,45 size 94x42; FormatPattern 9999
      ProcessValue <- "ST_FC_Var_g_N"
   TextField "Text Field_2" at 804,4 size 94x42; Text '产量kg / 篠送り出し速度 / 생산량kg'
   TextField "Text Field_24" at 899,4 size 94x42; Text '纱穗重量g / RunningMode / 運転モード / 코프중량'
   IOField "IO Field_4" at 804,45 size 94x42; FormatPattern 999.9
      ProcessValue <- "ST_Maintenance_HMI_r64_Production_Once"
   IOField "IO Field_5" at 899,46 size 94x42; FormatPattern 999.9
      ProcessValue <- "ST_Maintenance_HMI_r64_Weight_ShaSui"
   TextField "Text Field_3" at 614,4 size 94x42; Text '最大直径周期 / CarriageVelo / キャレージ速度 / 코프완성주기'
   IOField "IO Field_6" at 614,45 size 94x42; FormatPattern 9999
      ProcessValue <- "ST_FC_Var_g_ND"
   Button "OBJECT_106" at 1019,6 size 237x42; TextOff '手动 / EXIT'; TextList "mode_enabled_1"
      ProcessValue <- "ST_Main_Var_g_i16_Mode_Enabled"
      Appearance <- "ST_Main_Var_g_i16_Mode_Enabled"
   Button "OBJECT_111" at 1019,46 size 237x42; TextOff '手动 / EXIT'; TextList "automatic_status_1"
      Visibility <- "ST_Main_Var_g_bo_Mode_Enabled_Automatic"
      ProcessValue <- "ST_Main_Var_g_i16_Automatic_Status"
      Appearance <- "ST_Main_Var_g_i16_Automatic_Status"
   TextField "Text Field_40" at 234,4 size 94x42; Text '成纱支数'
   TextField "Text Field_43" at 329,4 size 94x42; Text '最大直径'
   TextField "Text Field_47" at 519,4 size 94x42; Text '单纱张力'
   TextField "Text Field_48" at 424,4 size 94x42; Text '纱穗个数'
   IOField "IO Field_69" at 234,45 size 94x42; FormatPattern 99.99
      ProcessValue <- "ST_HMI_Var_HMI_r64ZhiShu_ChengSha"
   IOField "IO Field_75" at 424,45 size 94x42; FormatPattern 9999
      ProcessValue <- "ST_HMI_Var_HMI_r64_ShuLiang_ShaSui"
   IOField "IO Field_76" at 519,45 size 94x42; FormatPattern 999.9
      ProcessValue <- "ST_HMI_Var_HMI_r64_LuoSha_Force_DanSha_ZhangLi_FangKai"
   IOField "IO Field_83" at 329,45 size 94x42; FormatPattern 99.9
      ProcessValue <- "ST_HMI_Var_HMI_r64Diameter_ShaSui_Max"
   Group "Group_电机温度" at 726,415 size 96x53
   Group "Group_驱动器温度" at 828,415 size 124x53
   Button "OBJECT_322" at 1152,493 size 119x60; TextOff '抬 弓 / EXIT'
      on Press: InvertBit("ST_MotionTask_ZhangLi_Var_HMI_bo_TaiGong")
      Appearance <- "ST_MotionTask_ZhangLi_Var_HMI_bo_TaiGong"
      ObjectEnable <- "ST_Main_Var_g_i16_Automatic_Status"
      Visibility <- "ST_Main_Var_g_i16_Automatic_Status"
   Group "Group_通用按钮" at 9,583 size 1262x60
   Button "OBJECT_9" at 1152,493 size 119x60; TextOff '抬 弓 / EXIT'
      on Press: InvertBit("ST_MotionTask_ZhangLi_Var_HMI_bo_TaiGong")
      Appearance <- "ST_MotionTask_ZhangLi_Var_HMI_bo_TaiGong"
      ObjectEnable <- "ST_Main_Var_g_i16_Automatic_Status"
      Visibility <- "ST_Main_Var_g_i16_Automatic_Status"
   Group "Group" at 9,493 size 445x60
   Group "Group_手动按钮隐藏" at 9,583 size 445x60
   TextField "Text Field_14" at 726,432 size 47x18; Text '锭子 / 番手: / 실 번수'
   TextField "Text Field_6" at 726,415 size 96x18; Text '电机温度(℃) / 番手: / 실 번수'
   TextField "Text Field_7" at 774,432 size 47x18; Text '张力 / 番手: / 실 번수'
   IOField "IO Field_15" at 726,450 size 47x18; FormatPattern 999.9
      ProcessValue <- "ST_Convert_ReadParameters_g_r64_SERVO_07_DingZi_35_Motor_temperature_real"
   IOField "IO Field_11" at 774,450 size 47x18; FormatPattern 999.9
      ProcessValue <- "ST_Convert_ReadParameters_g_r64_SERVO_04_ZhangLi_35_Motor_temperature_real"
   TextField "Text Field_8" at 828,432 size 61x18; Text '锭子 / 番手: / 실 번수'
   TextField "Text Field_10" at 890,432 size 61x18; Text '走车&张力 / 番手: / 실 번수'
   TextField "Text Field_9" at 828,415 size 124x18; Text '驱动器温度(℃) / 番手: / 실 번수'
   IOField "IO Field_19" at 828,450 size 61x18; FormatPattern 999.9
      ProcessValue <- "ST_Convert_ReadParameters_g_r64_SERVO_07_DingZi_37_4_Power_unit_temperatures_Interior_of_power_unit_real"
   IOField "IO Field_17" at 890,450 size 61x18; FormatPattern 999.9
      ProcessValue <- "ST_Convert_ReadParameters_g_r64_SERVO_03_ZouChe_37_4_Power_unit_temperatures_Interior_of_power_unit_real"
   Button "OBJECT_107" at 172,583 size 119x60; TextOff '手 动 / EXIT'
      on Release: ResetBit("ST_HMI_Var_HMI_bo_Manual")
      on Press: SetBit("ST_HMI_Var_HMI_bo_Manual")
      Appearance <- "ST_Main_Var_g_i16_Manual_Status"
   Button "OBJECT_108" at 498,583 size 119x60; TextOff '自 动 / EXIT'
      on Release: ResetBit("ST_HMI_Var_HMI_bo_Auto")
      on Press: SetBit("ST_HMI_Var_HMI_bo_Auto")
      Appearance <- "ST_Main_Var_g_bo_Mode_Enabled_Automatic"
   Button "OBJECT_109" at 662,583 size 119x60; TextOff '启 动 / EXIT'
      on Release: ResetBit("ST_HMI_Var_HMI_bo_ZiDong_QiDong")
      on Press: SetBit("ST_HMI_Var_HMI_bo_ZiDong_QiDong")
      Appearance <- "ST_Main_Var_g_bo_Automatic_Running_Status"
      Visibility <- "ST_Main_Var_g_i16_Mode_Enabled"
   Button "OBJECT_110" at 825,583 size 119x60; TextOff '停 止 / EXIT'
      on Release: ResetBit("ST_HMI_Var_HMI_bo_ZiDong_TingZhi")
      on Press: SetBit("ST_HMI_Var_HMI_bo_ZiDong_TingZhi")
      Appearance <- "ST_Main_Var_g_i16_Automatic_Stopping_Selected"
      Visibility <- "ST_Main_Var_g_bo_Mode_Enabled_Automatic"
   Button "OBJECT_117" at 988,583 size 119x60; TextOff '紧急停止 / EXIT'
      on Release: SetBit("ST_HMI_Var_HMI_bo_ZiDong_JiTing")
      on Press: ResetBit("ST_HMI_Var_HMI_bo_ZiDong_JiTing")
      Visibility <- "ST_Main_Var_g_i16_Mode_Enabled"
   Button "OBJECT_118" at 1152,583 size 119x60; TextOff '退出急停 / EXIT'
      on Press: SetTag("ST_Main_Var_g_i16_Automatic_Status", 1)
      Visibility <- "ST_Main_Var_g_bo_Automatic_Status_Mergestop"
   Button "OBJECT_1" at 9,583 size 119x60; TextOff '去使能 / EXIT'
      on Release: ResetBit("ST_HMI_Var_HMI_bo_Disable")
      on Press: SetBit("ST_HMI_Var_HMI_bo_Disable")
      Appearance <- "ST_Main_Var_g_i16_Disable_Status"
   Button "OBJECT_2" at 335,583 size 119x60; TextOff '回起点 / EXIT'
      on Release: ResetBit("ST_HMI_Var_HMI_bo_Start_Position")
      on Press: SetBit("ST_HMI_Var_HMI_bo_Start_Position")
      Appearance <- "ST_Main_Var_g_i16_Mode_Enabled"
   Group "Group_生头按钮" at 662,583 size 282x60
   Button "OBJECT_5" at 825,583 size 119x60; TextOff '停 止 / EXIT'
      on Release: ResetBit("ST_HMI_Var_HMI_bo_ShengTou_TingZhi")
      on Press: SetBit("ST_HMI_Var_HMI_bo_ShengTou_TingZhi")
      Visibility <- "ST_Main_Var_g_i16_Mode_Enabled"
      Appearance <- "ST_Main_Var_g_bo_KongDing_Running_Status"
   Button "OBJECT_4" at 662,583 size 119x60; TextOff '启 动 / EXIT'
      on Release: ResetBit("ST_HMI_Var_HMI_bo_ShengTou_QiDong")
      on Press: SetBit("ST_HMI_Var_HMI_bo_ShengTou_QiDong")
      Visibility <- "ST_Main_Var_g_i16_Mode_Enabled"
      Appearance <- "ST_Main_Var_g_bo_KongDing_Running_Status"
   Group "Group_抬弓设定" at 1040,169 size 189x127; Authorization "User administration"
   TextField "Text Field_12" at 1040,169 size 188x42; Text '抬弓设定'
      Visibility <- "ST_MotionTask_ZhangLi_Var_HMI_bo_TaiGong"
   TextField "Text Field_4" at 1135,211 size 94x42; Text '抬弓角度'
      Visibility <- "ST_MotionTask_ZhangLi_Var_HMI_bo_TaiGong"
   TextField "Text Field_5" at 1040,211 size 94x42; Text '放下位置'
      Visibility <- "ST_MotionTask_ZhangLi_Var_HMI_bo_TaiGong"
   IOField "IO Field_102" at 1135,254 size 94x42; Authorization "User administration"; FormatPattern 99
      Visibility <- "ST_MotionTask_ZhangLi_Var_HMI_bo_TaiGong"
      ProcessValue <- "ST_MotionTask_ZhangLi_Var_HMI_r64Axis_1_ZhangLi_Position_TaiGong"
   IOField "IO Field_101" at 1040,254 size 94x42; Authorization "User administration"; FormatPattern 9999
      Visibility <- "ST_MotionTask_ZhangLi_Var_HMI_bo_TaiGong"
      ProcessValue <- "ST_MotionTask_ZhangLi_Var_HMI_r64Axis_ZouChe_Position_TaiGong_FangXia"
   Line "线_211" at 1134,212 size 0x84
      Visibility <- "ST_MotionTask_ZhangLi_Var_HMI_bo_TaiGong"
   Rectangle "矩形_411" at 1152,493 size 119x60
      Visibility <- "ST_Main_Var_g_i16_Mode_Enabled"
   Group "Group_生头设定" at 1039,97 size 190x260
   TextField "Text Field_49" at 1040,182 size 94x42; Text '单纱张力'
      Visibility <- "ST_Main_Var_g_i16_Mode_Enabled"
   TextField "Text Field_52" at 1040,225 size 94x42; Text '弓目标值'
      Visibility <- "ST_Main_Var_g_i16_Mode_Enabled"
   IOField "IO Field_511" at 1135,182 size 94x42; FormatPattern 999.9
      Visibility <- "ST_Main_Var_g_i16_Mode_Enabled"
      ProcessValue <- "ST_HMI_Var_HMI_r64_DanSha_ZhangLi_ShengTou"
   IOField "IO Field_79" at 1135,225 size 94x42; FormatPattern 999.9
      Visibility <- "ST_Main_Var_g_i16_Mode_Enabled"
      ProcessValue <- "ST_HMI_Var_HMI_r64Axis_1_ZhangLi_Position_JuanRao_Set_KongDing_12"
   TextField "Text Field_62" at 1040,139 size 94x42; Text '出车展距:'
      Visibility <- "ST_Main_Var_g_i16_Mode_Enabled"
   IOField "IO Field_35" at 1135,139 size 94x42; FormatPattern 9999
      Visibility <- "ST_Main_Var_g_i16_Mode_Enabled"
      ProcessValue <- "ST_HMI_Var_HMI_r64Position_ChuChe_KongDing_7"
   TextField "Text Field_11" at 1040,97 size 189x42; Text '生头设定'
      Visibility <- "ST_Main_Var_g_i16_Mode_Enabled"
   Button "OBJECT_7" at 1039,315 size 94x42; TextOff '纱管1 / EXIT'; Authorization "Monitor"
      on Press: SetTag("ST_HMI_Var_HMI_i16_Status_ShaGuan_Select", 1)
      Appearance <- "ST_HMI_Var_HMI_i16_Status_ShaGuan_Select"
      Visibility <- "ST_Main_Var_g_i16_Mode_Enabled"
   Button "OBJECT_8" at 1134,315 size 94x42; TextOff '纱管2 / EXIT'; Authorization "Monitor"
      on Press: SetTag("ST_HMI_Var_HMI_i16_Status_ShaGuan_Select", 2)
      Appearance <- "ST_HMI_Var_HMI_i16_Status_ShaGuan_Select"
      Visibility <- "ST_Main_Var_g_i16_Mode_Enabled"
   TextField "Text Field_13" at 1040,268 size 94x42; Text '速度比例'
      Visibility <- "ST_Main_Var_g_i16_Mode_Enabled"
   IOField "IO Field_519" at 1135,268 size 94x42; FormatPattern 9.99
      Visibility <- "ST_Main_Var_g_i16_Mode_Enabled"
      ProcessValue <- "ST_HMI_Var_HMI_r64_Scale_KongDing_7"
   Button "OBJECT_3" at 9,493 size 119x60; TextOff '空锭(插管) / EXIT'
      on Release: ResetBit("ST_HMI_Var_HMI_bo_KongDingShengTou")
      on Press: SetBit("ST_HMI_Var_HMI_bo_KongDingShengTou")
      Appearance <- "ST_HMI_Var_HMI_i16_ShengTou_Select"
      Visibility <- "ST_Main_Var_g_i16_Mode_Enabled"
   Button "OBJECT_312" at 335,493 size 119x60; TextOff '落纱生头 / EXIT'
      on Release: ResetBit("ST_HMI_Var_HMI_bo_LuoShaShengTou")
      on Press: SetBit("ST_HMI_Var_HMI_bo_LuoShaShengTou")
      Appearance <- "ST_HMI_Var_HMI_i16_ShengTou_Select"
      Visibility <- "ST_Main_Var_g_i16_Mode_Enabled"
   Button "OBJECT_6" at 172,493 size 119x60; TextOff '空锭(光锭) / EXIT'
      on Release: ResetBit("ST_HMI_Var_HMI_bo_KongDingShengTou_GuangDing")
      on Press: SetBit("ST_HMI_Var_HMI_bo_KongDingShengTou_GuangDing")
      Appearance <- "ST_HMI_Var_HMI_i16_ShengTou_Select"
      Visibility <- "ST_Main_Var_g_i16_Mode_Enabled"
   Rectangle "手动按钮隐藏_3" at 9,583 size 119x60
      Visibility <- "ST_Main_Var_g_bo_Automatic_Running_Status"
   Rectangle "手动按钮隐藏_2" at 172,583 size 119x60
      Visibility <- "ST_Main_Var_g_bo_Automatic_Running_Status"
   Rectangle "手动按钮隐藏_1" at 335,583 size 119x60
      Visibility <- "ST_Main_Var_g_bo_Automatic_Running_Status"

